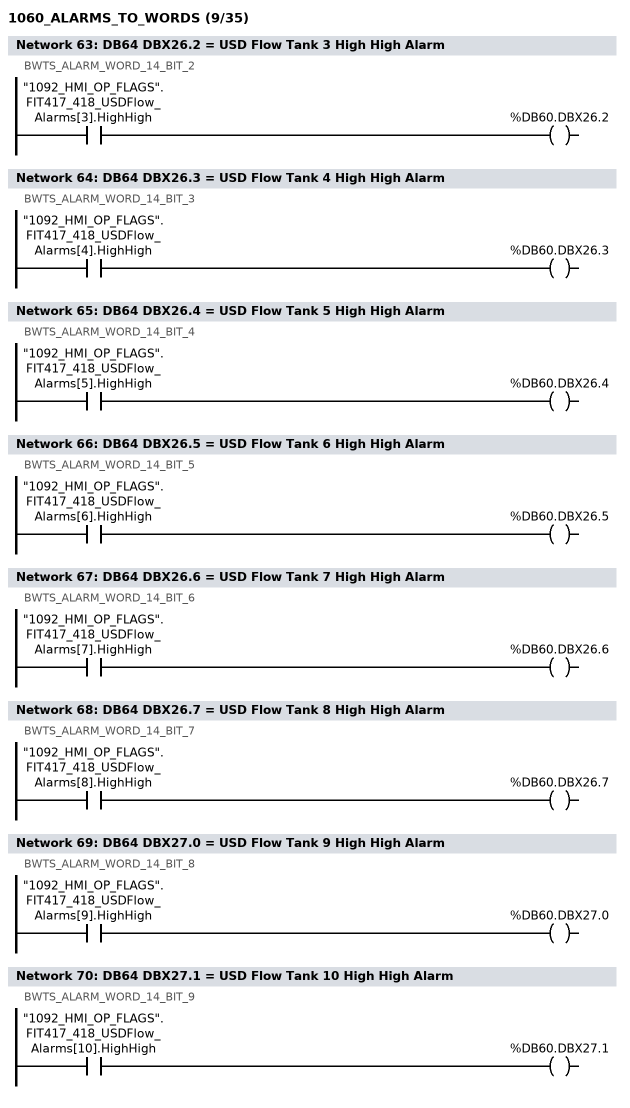
   RUNG wire#powerrail
      Contact( "1092_HMI_OP_FLAGS".FIT417_418_USDFlow_Alarms[3].HighHigh )
      Coil( %DB60.DBX26.2 )
   END_RUNG
   // the same network as SCL:
   %DB60.DBX26.2 := "1092_HMI_OP_FLAGS".FIT417_418_USDFlow_Alarms[3].HighHigh;
END_REGION

REGION Network 64: DB64 DBX26.3 = USD Flow Tank 4 High High Alarm
   // BWTS_ALARM_WORD_14_BIT_3
   RUNG wire#powerrail
      Contact( "1092_HMI_OP_FLAGS".FIT417_418_USDFlow_Alarms[4].HighHigh )
      Coil( %DB60.DBX26.3 )
   END_RUNG
   // the same network as SCL:
   %DB60.DBX26.3 := "1092_HMI_OP_FLAGS".FIT417_418_USDFlow_Alarms[4].HighHigh;
END_REGION

REGION Network 65: DB64 DBX26.4 = USD Flow Tank 5 High High Alarm
   // BWTS_ALARM_WORD_14_BIT_4
   RUNG wire#powerrail
      Contact( "1092_HMI_OP_FLAGS".FIT417_418_USDFlow_Alarms[5].HighHigh )
      Coil( %DB60.DBX26.4 )
   END_RUNG
   // the same network as SCL:
   %DB60.DBX26.4 := "1092_HMI_OP_FLAGS".FIT417_418_USDFlow_Alarms[5].HighHigh;
END_REGION

REGION Network 66: DB64 DBX26.5 = USD Flow Tank 6 High High Alarm
   // BWTS_ALARM_WORD_14_BIT_5
   RUNG wire#powerrail
      Contact( "1092_HMI_OP_FLAGS".FIT417_418_USDFlow_Alarms[6].HighHigh )
      Coil( %DB60.DBX26.5 )
   END_RUNG
   // the same network as SCL:
   %DB60.DBX26.5 := "1092_HMI_OP_FLAGS".FIT417_418_USDFlow_Alarms[6].HighHigh;
END_REGION

REGION Network 67: DB64 DBX26.6 = USD Flow Tank 7 High High Alarm
   // BWTS_ALARM_WORD_14_BIT_6
   RUNG wire#powerrail
      Contact( "1092_HMI_OP_FLAGS".FIT417_418_USDFlow_Alarms[7].HighHigh )
      Coil( %DB60.DBX26.6 )
   END_RUNG
   // the same network as SCL:
   %DB60.DBX26.6 := "1092_HMI_OP_FLAGS".FIT417_418_USDFlow_Alarms[7].HighHigh;
END_REGION

REGION Network 68: DB64 DBX26.7 = USD Flow Tank 8 High High Alarm
   // BWTS_ALARM_WORD_14_BIT_7
   RUNG wire#powerrail
      Contact( "1092_HMI_OP_FLAGS".FIT417_418_USDFlow_Alarms[8].HighHigh )
      Coil( %DB60.DBX26.7 )
   END_RUNG
   // the same network as SCL:
   %DB60.DBX26.7 := "1092_HMI_OP_FLAGS".FIT417_418_USDFlow_Alarms[8].HighHigh;
END_REGION

REGION Network 69: DB64 DBX27.0 = USD Flow Tank 9 High High Alarm
   // BWTS_ALARM_WORD_14_BIT_8
   RUNG wire#powerrail
      Contact( "1092_HMI_OP_FLAGS".FIT417_418_USDFlow_Alarms[9].HighHigh )
      Coil( %DB60.DBX27.0 )
   END_RUNG
   // the same network as SCL:
   %DB60.DBX27.0 := "1092_HMI_OP_FLAGS".FIT417_418_USDFlow_Alarms[9].HighHigh;
END_REGION

REGION Network 70: DB64 DBX27.1 = USD Flow Tank 10 High High Alarm
   // BWTS_ALARM_WORD_14_BIT_9
   RUNG wire#powerrail
      Contact( "1092_HMI_OP_FLAGS".FIT417_418_USDFlow_Alarms[10].HighHigh )
      Coil( %DB60.DBX27.1 )
   END_RUNG
   // the same network as SCL:
   %DB60.DBX27.1 := "1092_HMI_OP_FLAGS".FIT417_418_USDFlow_Alarms[10].HighHigh;
END_REGION

REGION Network 71: DB64 DBX27.2 = USD Flow Tank 11 High High Alarm
   // BWTS_ALARM_WORD_14_BIT_10
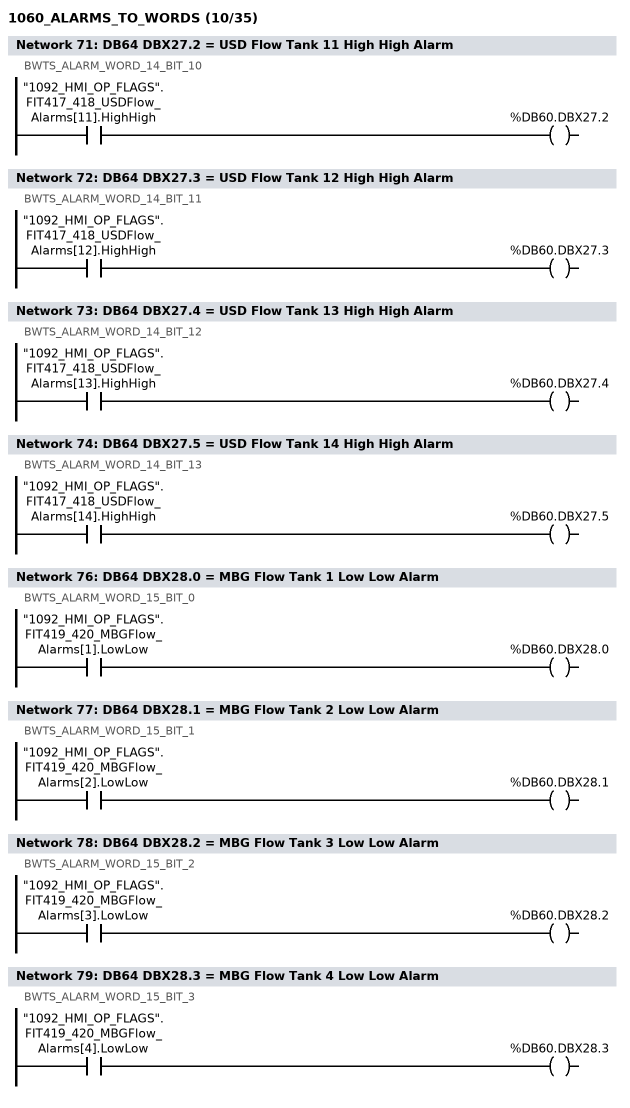
   RUNG wire#powerrail
      Contact( "1092_HMI_OP_FLAGS".FIT417_418_USDFlow_Alarms[11].HighHigh )
      Coil( %DB60.DBX27.2 )
   END_RUNG
   // the same network as SCL:
   %DB60.DBX27.2 := "1092_HMI_OP_FLAGS".FIT417_418_USDFlow_Alarms[11].HighHigh;
END_REGION

REGION Network 72: DB64 DBX27.3 = USD Flow Tank 12 High High Alarm
   // BWTS_ALARM_WORD_14_BIT_11
   RUNG wire#powerrail
      Contact( "1092_HMI_OP_FLAGS".FIT417_418_USDFlow_Alarms[12].HighHigh )
      Coil( %DB60.DBX27.3 )
   END_RUNG
   // the same network as SCL:
   %DB60.DBX27.3 := "1092_HMI_OP_FLAGS".FIT417_418_USDFlow_Alarms[12].HighHigh;
END_REGION

REGION Network 73: DB64 DBX27.4 = USD Flow Tank 13 High High Alarm
   // BWTS_ALARM_WORD_14_BIT_12
   RUNG wire#powerrail
      Contact( "1092_HMI_OP_FLAGS".FIT417_418_USDFlow_Alarms[13].HighHigh )
      Coil( %DB60.DBX27.4 )
   END_RUNG
   // the same network as SCL:
   %DB60.DBX27.4 := "1092_HMI_OP_FLAGS".FIT417_418_USDFlow_Alarms[13].HighHigh;
END_REGION

REGION Network 74: DB64 DBX27.5 = USD Flow Tank 14 High High Alarm
   // BWTS_ALARM_WORD_14_BIT_13
   RUNG wire#powerrail
      Contact( "1092_HMI_OP_FLAGS".FIT417_418_USDFlow_Alarms[14].HighHigh )
      Coil( %DB60.DBX27.5 )
   END_RUNG
   // the same network as SCL:
   %DB60.DBX27.5 := "1092_HMI_OP_FLAGS".FIT417_418_USDFlow_Alarms[14].HighHigh;
END_REGION

REGION Network 76: DB64 DBX28.0 = MBG Flow Tank 1 Low Low Alarm
   // BWTS_ALARM_WORD_15_BIT_0
   RUNG wire#powerrail
      Contact( "1092_HMI_OP_FLAGS".FIT419_420_MBGFlow_Alarms[1].LowLow )
      Coil( %DB60.DBX28.0 )
   END_RUNG
   // the same network as SCL:
   %DB60.DBX28.0 := "1092_HMI_OP_FLAGS".FIT419_420_MBGFlow_Alarms[1].LowLow;
END_REGION

REGION Network 77: DB64 DBX28.1 = MBG Flow Tank 2 Low Low Alarm
   // BWTS_ALARM_WORD_15_BIT_1
   RUNG wire#powerrail
      Contact( "1092_HMI_OP_FLAGS".FIT419_420_MBGFlow_Alarms[2].LowLow )
      Coil( %DB60.DBX28.1 )
   END_RUNG
   // the same network as SCL:
   %DB60.DBX28.1 := "1092_HMI_OP_FLAGS".FIT419_420_MBGFlow_Alarms[2].LowLow;
END_REGION

REGION Network 78: DB64 DBX28.2 = MBG Flow Tank 3 Low Low Alarm
   // BWTS_ALARM_WORD_15_BIT_2
   RUNG wire#powerrail
      Contact( "1092_HMI_OP_FLAGS".FIT419_420_MBGFlow_Alarms[3].LowLow )
      Coil( %DB60.DBX28.2 )
   END_RUNG
   // the same network as SCL:
   %DB60.DBX28.2 := "1092_HMI_OP_FLAGS".FIT419_420_MBGFlow_Alarms[3].LowLow;
END_REGION

REGION Network 79: DB64 DBX28.3 = MBG Flow Tank 4 Low Low Alarm
   // BWTS_ALARM_WORD_15_BIT_3
   RUNG wire#powerrail
      Contact( "1092_HMI_OP_FLAGS".FIT419_420_MBGFlow_Alarms[4].LowLow )
      Coil( %DB60.DBX28.3 )
   END_RUNG
   // the same network as SCL:
   %DB60.DBX28.3 := "1092_HMI_OP_FLAGS".FIT419_420_MBGFlow_Alarms[4].LowLow;
END_REGION

REGION Network 80: DB64 DBX28.4 = MBG Flow Tank 5 Low Low Alarm
   // BWTS_ALARM_WORD_15_BIT_4
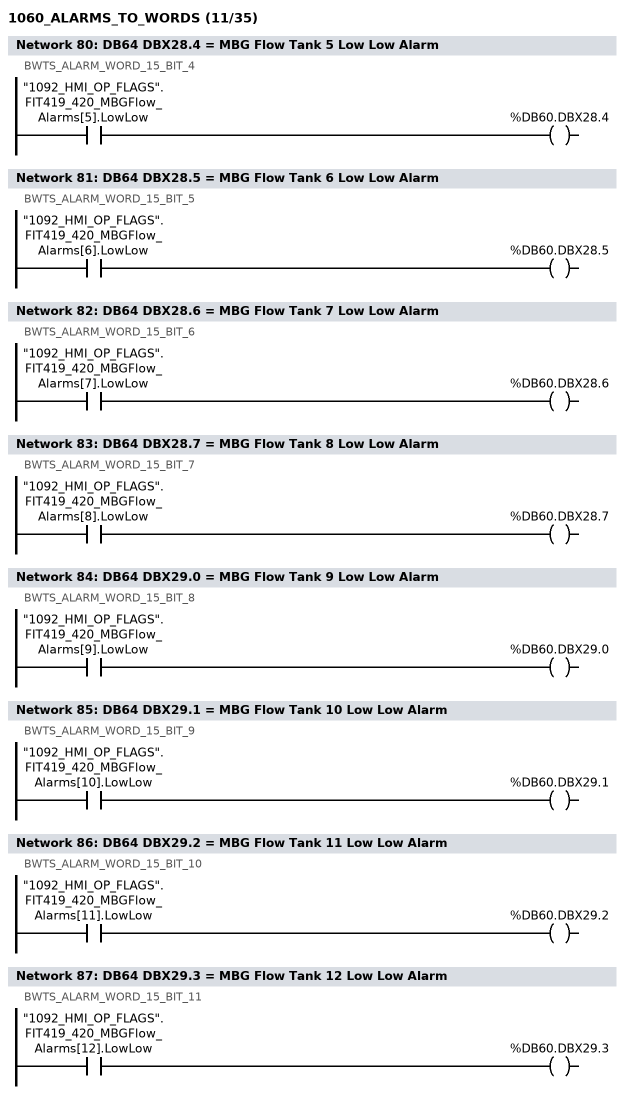
   RUNG wire#powerrail
      Contact( "1092_HMI_OP_FLAGS".FIT419_420_MBGFlow_Alarms[5].LowLow )
      Coil( %DB60.DBX28.4 )
   END_RUNG
   // the same network as SCL:
   %DB60.DBX28.4 := "1092_HMI_OP_FLAGS".FIT419_420_MBGFlow_Alarms[5].LowLow;
END_REGION

REGION Network 81: DB64 DBX28.5 = MBG Flow Tank 6 Low Low Alarm
   // BWTS_ALARM_WORD_15_BIT_5
   RUNG wire#powerrail
      Contact( "1092_HMI_OP_FLAGS".FIT419_420_MBGFlow_Alarms[6].LowLow )
      Coil( %DB60.DBX28.5 )
   END_RUNG
   // the same network as SCL:
   %DB60.DBX28.5 := "1092_HMI_OP_FLAGS".FIT419_420_MBGFlow_Alarms[6].LowLow;
END_REGION

REGION Network 82: DB64 DBX28.6 = MBG Flow Tank 7 Low Low Alarm
   // BWTS_ALARM_WORD_15_BIT_6
   RUNG wire#powerrail
      Contact( "1092_HMI_OP_FLAGS".FIT419_420_MBGFlow_Alarms[7].LowLow )
      Coil( %DB60.DBX28.6 )
   END_RUNG
   // the same network as SCL:
   %DB60.DBX28.6 := "1092_HMI_OP_FLAGS".FIT419_420_MBGFlow_Alarms[7].LowLow;
END_REGION

REGION Network 83: DB64 DBX28.7 = MBG Flow Tank 8 Low Low Alarm
   // BWTS_ALARM_WORD_15_BIT_7
   RUNG wire#powerrail
      Contact( "1092_HMI_OP_FLAGS".FIT419_420_MBGFlow_Alarms[8].LowLow )
      Coil( %DB60.DBX28.7 )
   END_RUNG
   // the same network as SCL:
   %DB60.DBX28.7 := "1092_HMI_OP_FLAGS".FIT419_420_MBGFlow_Alarms[8].LowLow;
END_REGION

REGION Network 84: DB64 DBX29.0 = MBG Flow Tank 9 Low Low Alarm
   // BWTS_ALARM_WORD_15_BIT_8
   RUNG wire#powerrail
      Contact( "1092_HMI_OP_FLAGS".FIT419_420_MBGFlow_Alarms[9].LowLow )
      Coil( %DB60.DBX29.0 )
   END_RUNG
   // the same network as SCL:
   %DB60.DBX29.0 := "1092_HMI_OP_FLAGS".FIT419_420_MBGFlow_Alarms[9].LowLow;
END_REGION

REGION Network 85: DB64 DBX29.1 = MBG Flow Tank 10 Low Low Alarm
   // BWTS_ALARM_WORD_15_BIT_9
   RUNG wire#powerrail
      Contact( "1092_HMI_OP_FLAGS".FIT419_420_MBGFlow_Alarms[10].LowLow )
      Coil( %DB60.DBX29.1 )
   END_RUNG
   // the same network as SCL:
   %DB60.DBX29.1 := "1092_HMI_OP_FLAGS".FIT419_420_MBGFlow_Alarms[10].LowLow;
END_REGION

REGION Network 86: DB64 DBX29.2 = MBG Flow Tank 11 Low Low Alarm
   // BWTS_ALARM_WORD_15_BIT_10
   RUNG wire#powerrail
      Contact( "1092_HMI_OP_FLAGS".FIT419_420_MBGFlow_Alarms[11].LowLow )
      Coil( %DB60.DBX29.2 )
   END_RUNG
   // the same network as SCL:
   %DB60.DBX29.2 := "1092_HMI_OP_FLAGS".FIT419_420_MBGFlow_Alarms[11].LowLow;
END_REGION

REGION Network 87: DB64 DBX29.3 = MBG Flow Tank 12 Low Low Alarm
   // BWTS_ALARM_WORD_15_BIT_11
   RUNG wire#powerrail
      Contact( "1092_HMI_OP_FLAGS".FIT419_420_MBGFlow_Alarms[12].LowLow )
      Coil( %DB60.DBX29.3 )
   END_RUNG
   // the same network as SCL:
   %DB60.DBX29.3 := "1092_HMI_OP_FLAGS".FIT419_420_MBGFlow_Alarms[12].LowLow;
END_REGION

REGION Network 88: DB64 DBX29.4 = MBG Flow Tank 13 Low Low Alarm
   // BWTS_ALARM_WORD_15_BIT_12
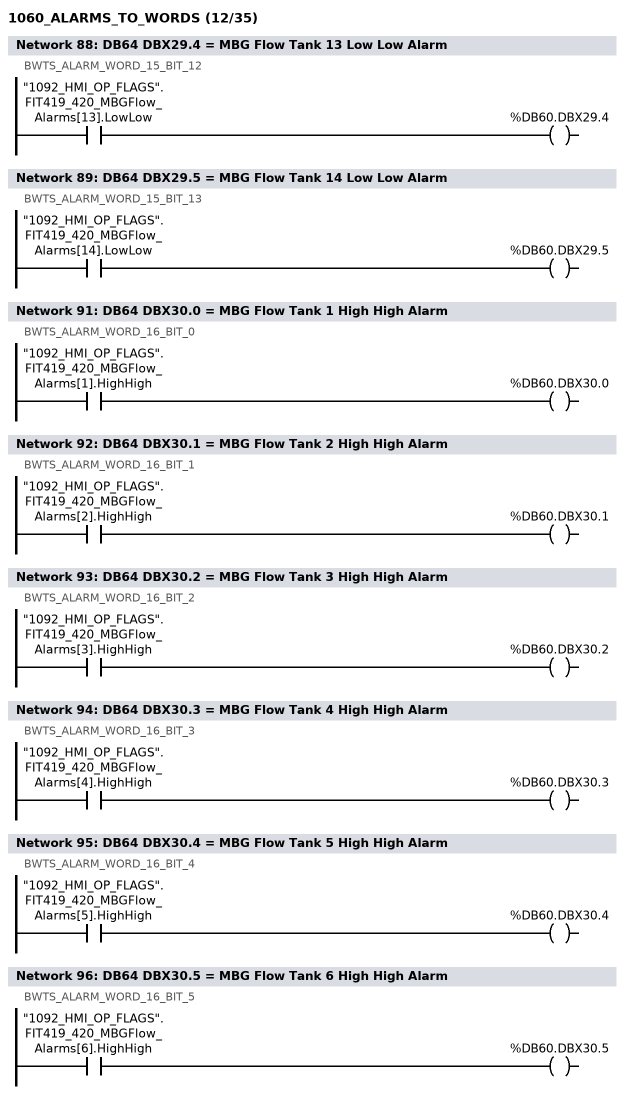
   RUNG wire#powerrail
      Contact( "1092_HMI_OP_FLAGS".FIT419_420_MBGFlow_Alarms[13].LowLow )
      Coil( %DB60.DBX29.4 )
   END_RUNG
   // the same network as SCL:
   %DB60.DBX29.4 := "1092_HMI_OP_FLAGS".FIT419_420_MBGFlow_Alarms[13].LowLow;
END_REGION

REGION Network 89: DB64 DBX29.5 = MBG Flow Tank 14 Low Low Alarm
   // BWTS_ALARM_WORD_15_BIT_13
   RUNG wire#powerrail
      Contact( "1092_HMI_OP_FLAGS".FIT419_420_MBGFlow_Alarms[14].LowLow )
      Coil( %DB60.DBX29.5 )
   END_RUNG
   // the same network as SCL:
   %DB60.DBX29.5 := "1092_HMI_OP_FLAGS".FIT419_420_MBGFlow_Alarms[14].LowLow;
END_REGION

REGION Network 91: DB64 DBX30.0 = MBG Flow Tank 1 High High Alarm
   // BWTS_ALARM_WORD_16_BIT_0
   RUNG wire#powerrail
      Contact( "1092_HMI_OP_FLAGS".FIT419_420_MBGFlow_Alarms[1].HighHigh )
      Coil( %DB60.DBX30.0 )
   END_RUNG
   // the same network as SCL:
   %DB60.DBX30.0 := "1092_HMI_OP_FLAGS".FIT419_420_MBGFlow_Alarms[1].HighHigh;
END_REGION

REGION Network 92: DB64 DBX30.1 = MBG Flow Tank 2 High High Alarm
   // BWTS_ALARM_WORD_16_BIT_1
   RUNG wire#powerrail
      Contact( "1092_HMI_OP_FLAGS".FIT419_420_MBGFlow_Alarms[2].HighHigh )
      Coil( %DB60.DBX30.1 )
   END_RUNG
   // the same network as SCL:
   %DB60.DBX30.1 := "1092_HMI_OP_FLAGS".FIT419_420_MBGFlow_Alarms[2].HighHigh;
END_REGION

REGION Network 93: DB64 DBX30.2 = MBG Flow Tank 3 High High Alarm
   // BWTS_ALARM_WORD_16_BIT_2
   RUNG wire#powerrail
      Contact( "1092_HMI_OP_FLAGS".FIT419_420_MBGFlow_Alarms[3].HighHigh )
      Coil( %DB60.DBX30.2 )
   END_RUNG
   // the same network as SCL:
   %DB60.DBX30.2 := "1092_HMI_OP_FLAGS".FIT419_420_MBGFlow_Alarms[3].HighHigh;
END_REGION

REGION Network 94: DB64 DBX30.3 = MBG Flow Tank 4 High High Alarm
   // BWTS_ALARM_WORD_16_BIT_3
   RUNG wire#powerrail
      Contact( "1092_HMI_OP_FLAGS".FIT419_420_MBGFlow_Alarms[4].HighHigh )
      Coil( %DB60.DBX30.3 )
   END_RUNG
   // the same network as SCL:
   %DB60.DBX30.3 := "1092_HMI_OP_FLAGS".FIT419_420_MBGFlow_Alarms[4].HighHigh;
END_REGION

REGION Network 95: DB64 DBX30.4 = MBG Flow Tank 5 High High Alarm
   // BWTS_ALARM_WORD_16_BIT_4
   RUNG wire#powerrail
      Contact( "1092_HMI_OP_FLAGS".FIT419_420_MBGFlow_Alarms[5].HighHigh )
      Coil( %DB60.DBX30.4 )
   END_RUNG
   // the same network as SCL:
   %DB60.DBX30.4 := "1092_HMI_OP_FLAGS".FIT419_420_MBGFlow_Alarms[5].HighHigh;
END_REGION

REGION Network 96: DB64 DBX30.5 = MBG Flow Tank 6 High High Alarm
   // BWTS_ALARM_WORD_16_BIT_5
   RUNG wire#powerrail
      Contact( "1092_HMI_OP_FLAGS".FIT419_420_MBGFlow_Alarms[6].HighHigh )
      Coil( %DB60.DBX30.5 )
   END_RUNG
   // the same network as SCL:
   %DB60.DBX30.5 := "1092_HMI_OP_FLAGS".FIT419_420_MBGFlow_Alarms[6].HighHigh;
END_REGION

REGION Network 97: DB64 DBX30.6 = MBG Flow Tank 7 High High Alarm
   // BWTS_ALARM_WORD_16_BIT_6
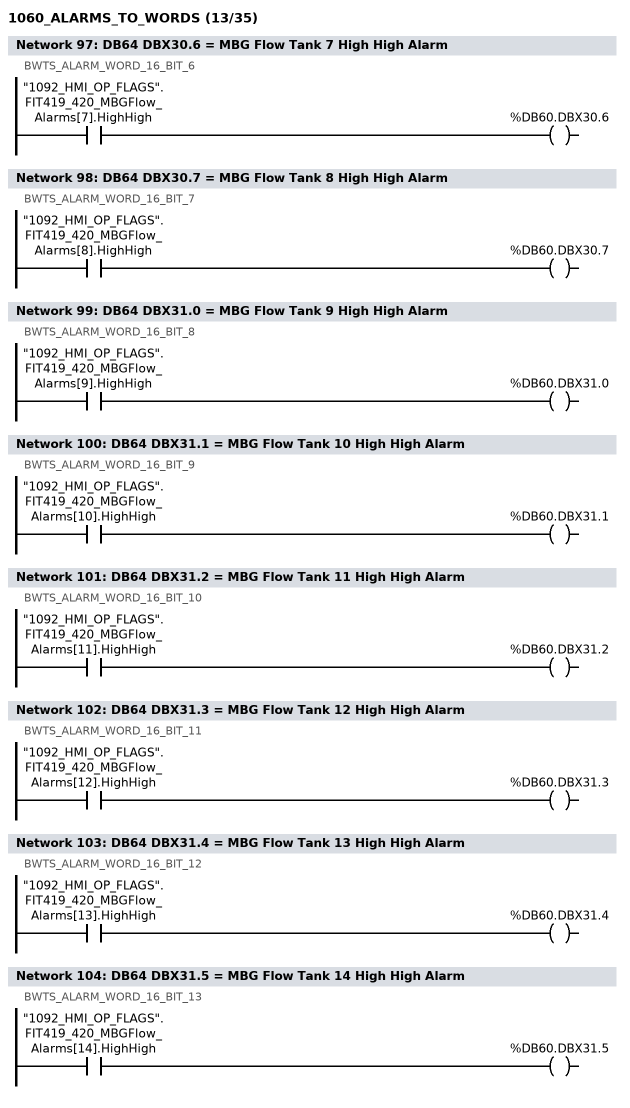
   RUNG wire#powerrail
      Contact( "1092_HMI_OP_FLAGS".FIT419_420_MBGFlow_Alarms[7].HighHigh )
      Coil( %DB60.DBX30.6 )
   END_RUNG
   // the same network as SCL:
   %DB60.DBX30.6 := "1092_HMI_OP_FLAGS".FIT419_420_MBGFlow_Alarms[7].HighHigh;
END_REGION

REGION Network 98: DB64 DBX30.7 = MBG Flow Tank 8 High High Alarm
   // BWTS_ALARM_WORD_16_BIT_7
   RUNG wire#powerrail
      Contact( "1092_HMI_OP_FLAGS".FIT419_420_MBGFlow_Alarms[8].HighHigh )
      Coil( %DB60.DBX30.7 )
   END_RUNG
   // the same network as SCL:
   %DB60.DBX30.7 := "1092_HMI_OP_FLAGS".FIT419_420_MBGFlow_Alarms[8].HighHigh;
END_REGION

REGION Network 99: DB64 DBX31.0 = MBG Flow Tank 9 High High Alarm
   // BWTS_ALARM_WORD_16_BIT_8
   RUNG wire#powerrail
      Contact( "1092_HMI_OP_FLAGS".FIT419_420_MBGFlow_Alarms[9].HighHigh )
      Coil( %DB60.DBX31.0 )
   END_RUNG
   // the same network as SCL:
   %DB60.DBX31.0 := "1092_HMI_OP_FLAGS".FIT419_420_MBGFlow_Alarms[9].HighHigh;
END_REGION

REGION Network 100: DB64 DBX31.1 = MBG Flow Tank 10 High High Alarm
   // BWTS_ALARM_WORD_16_BIT_9
   RUNG wire#powerrail
      Contact( "1092_HMI_OP_FLAGS".FIT419_420_MBGFlow_Alarms[10].HighHigh )
      Coil( %DB60.DBX31.1 )
   END_RUNG
   // the same network as SCL:
   %DB60.DBX31.1 := "1092_HMI_OP_FLAGS".FIT419_420_MBGFlow_Alarms[10].HighHigh;
END_REGION

REGION Network 101: DB64 DBX31.2 = MBG Flow Tank 11 High High Alarm
   // BWTS_ALARM_WORD_16_BIT_10
   RUNG wire#powerrail
      Contact( "1092_HMI_OP_FLAGS".FIT419_420_MBGFlow_Alarms[11].HighHigh )
      Coil( %DB60.DBX31.2 )
   END_RUNG
   // the same network as SCL:
   %DB60.DBX31.2 := "1092_HMI_OP_FLAGS".FIT419_420_MBGFlow_Alarms[11].HighHigh;
END_REGION

REGION Network 102: DB64 DBX31.3 = MBG Flow Tank 12 High High Alarm
   // BWTS_ALARM_WORD_16_BIT_11
   RUNG wire#powerrail
      Contact( "1092_HMI_OP_FLAGS".FIT419_420_MBGFlow_Alarms[12].HighHigh )
      Coil( %DB60.DBX31.3 )
   END_RUNG
   // the same network as SCL:
   %DB60.DBX31.3 := "1092_HMI_OP_FLAGS".FIT419_420_MBGFlow_Alarms[12].HighHigh;
END_REGION

REGION Network 103: DB64 DBX31.4 = MBG Flow Tank 13 High High Alarm
   // BWTS_ALARM_WORD_16_BIT_12
   RUNG wire#powerrail
      Contact( "1092_HMI_OP_FLAGS".FIT419_420_MBGFlow_Alarms[13].HighHigh )
      Coil( %DB60.DBX31.4 )
   END_RUNG
   // the same network as SCL:
   %DB60.DBX31.4 := "1092_HMI_OP_FLAGS".FIT419_420_MBGFlow_Alarms[13].HighHigh;
END_REGION

REGION Network 104: DB64 DBX31.5 = MBG Flow Tank 14 High High Alarm
   // BWTS_ALARM_WORD_16_BIT_13
   RUNG wire#powerrail
      Contact( "1092_HMI_OP_FLAGS".FIT419_420_MBGFlow_Alarms[14].HighHigh )
      Coil( %DB60.DBX31.5 )
   END_RUNG
   // the same network as SCL:
   %DB60.DBX31.5 := "1092_HMI_OP_FLAGS".FIT419_420_MBGFlow_Alarms[14].HighHigh;
END_REGION

REGION Network 106: DB64 DBX32.0 = BWT Level Tank 1 Low Alarm
   // BWTS_ALARM_WORD_17_BIT_0
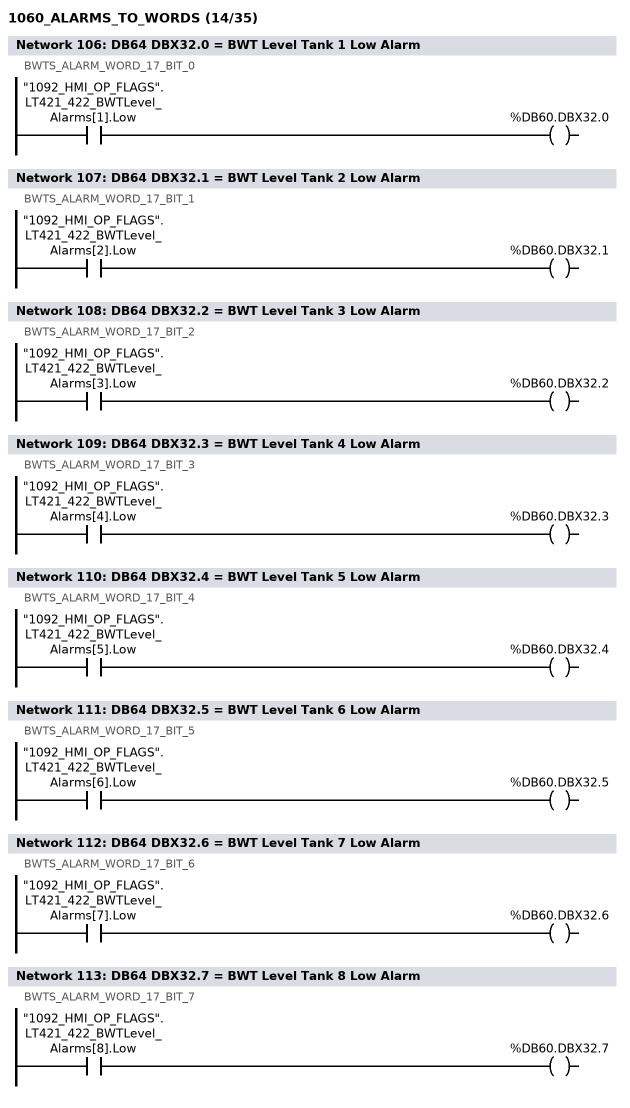
   RUNG wire#powerrail
      Contact( "1092_HMI_OP_FLAGS".LT421_422_BWTLevel_Alarms[1].Low )
      Coil( %DB60.DBX32.0 )
   END_RUNG
   // the same network as SCL:
   %DB60.DBX32.0 := "1092_HMI_OP_FLAGS".LT421_422_BWTLevel_Alarms[1].Low;
END_REGION

REGION Network 107: DB64 DBX32.1 = BWT Level Tank 2 Low Alarm
   // BWTS_ALARM_WORD_17_BIT_1
   RUNG wire#powerrail
      Contact( "1092_HMI_OP_FLAGS".LT421_422_BWTLevel_Alarms[2].Low )
      Coil( %DB60.DBX32.1 )
   END_RUNG
   // the same network as SCL:
   %DB60.DBX32.1 := "1092_HMI_OP_FLAGS".LT421_422_BWTLevel_Alarms[2].Low;
END_REGION

REGION Network 108: DB64 DBX32.2 = BWT Level Tank 3 Low Alarm
   // BWTS_ALARM_WORD_17_BIT_2
   RUNG wire#powerrail
      Contact( "1092_HMI_OP_FLAGS".LT421_422_BWTLevel_Alarms[3].Low )
      Coil( %DB60.DBX32.2 )
   END_RUNG
   // the same network as SCL:
   %DB60.DBX32.2 := "1092_HMI_OP_FLAGS".LT421_422_BWTLevel_Alarms[3].Low;
END_REGION

REGION Network 109: DB64 DBX32.3 = BWT Level Tank 4 Low Alarm
   // BWTS_ALARM_WORD_17_BIT_3
   RUNG wire#powerrail
      Contact( "1092_HMI_OP_FLAGS".LT421_422_BWTLevel_Alarms[4].Low )
      Coil( %DB60.DBX32.3 )
   END_RUNG
   // the same network as SCL:
   %DB60.DBX32.3 := "1092_HMI_OP_FLAGS".LT421_422_BWTLevel_Alarms[4].Low;
END_REGION

REGION Network 110: DB64 DBX32.4 = BWT Level Tank 5 Low Alarm
   // BWTS_ALARM_WORD_17_BIT_4
   RUNG wire#powerrail
      Contact( "1092_HMI_OP_FLAGS".LT421_422_BWTLevel_Alarms[5].Low )
      Coil( %DB60.DBX32.4 )
   END_RUNG
   // the same network as SCL:
   %DB60.DBX32.4 := "1092_HMI_OP_FLAGS".LT421_422_BWTLevel_Alarms[5].Low;
END_REGION

REGION Network 111: DB64 DBX32.5 = BWT Level Tank 6 Low Alarm
   // BWTS_ALARM_WORD_17_BIT_5
   RUNG wire#powerrail
      Contact( "1092_HMI_OP_FLAGS".LT421_422_BWTLevel_Alarms[6].Low )
      Coil( %DB60.DBX32.5 )
   END_RUNG
   // the same network as SCL:
   %DB60.DBX32.5 := "1092_HMI_OP_FLAGS".LT421_422_BWTLevel_Alarms[6].Low;
END_REGION

REGION Network 112: DB64 DBX32.6 = BWT Level Tank 7 Low Alarm
   // BWTS_ALARM_WORD_17_BIT_6
   RUNG wire#powerrail
      Contact( "1092_HMI_OP_FLAGS".LT421_422_BWTLevel_Alarms[7].Low )
      Coil( %DB60.DBX32.6 )
   END_RUNG
   // the same network as SCL:
   %DB60.DBX32.6 := "1092_HMI_OP_FLAGS".LT421_422_BWTLevel_Alarms[7].Low;
END_REGION

REGION Network 113: DB64 DBX32.7 = BWT Level Tank 8 Low Alarm
   // BWTS_ALARM_WORD_17_BIT_7
   RUNG wire#powerrail
      Contact( "1092_HMI_OP_FLAGS".LT421_422_BWTLevel_Alarms[8].Low )
      Coil( %DB60.DBX32.7 )
   END_RUNG
   // the same network as SCL:
   %DB60.DBX32.7 := "1092_HMI_OP_FLAGS".LT421_422_BWTLevel_Alarms[8].Low;
END_REGION

REGION Network 114: DB64 DBX33.0 = BWT Level Tank 9 Low Alarm
   // BWTS_ALARM_WORD_17_BIT_8
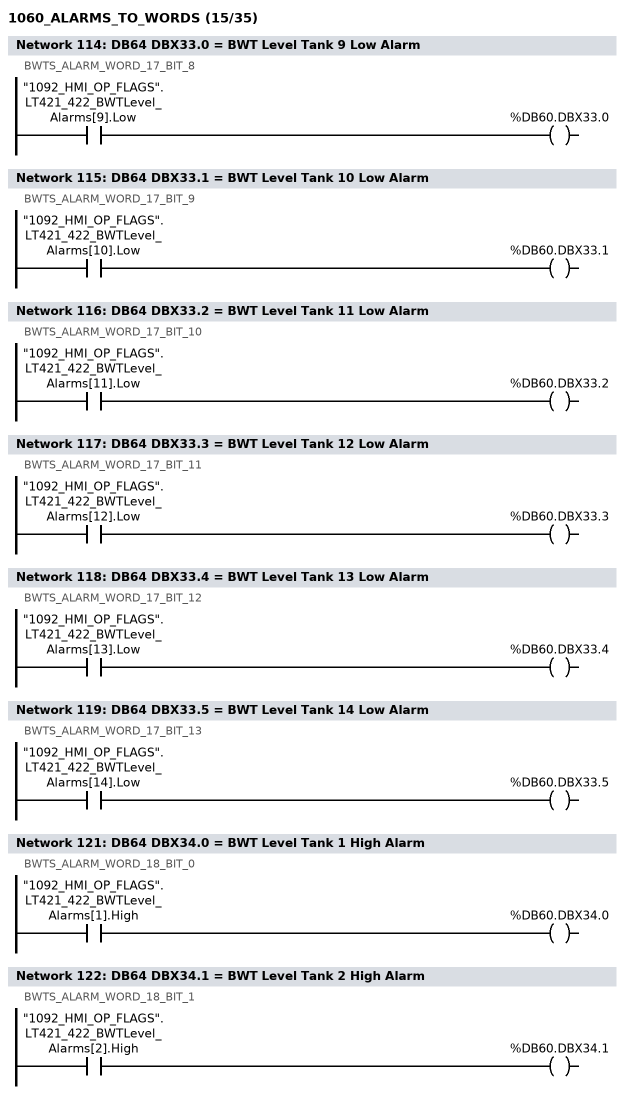
   RUNG wire#powerrail
      Contact( "1092_HMI_OP_FLAGS".LT421_422_BWTLevel_Alarms[9].Low )
      Coil( %DB60.DBX33.0 )
   END_RUNG
   // the same network as SCL:
   %DB60.DBX33.0 := "1092_HMI_OP_FLAGS".LT421_422_BWTLevel_Alarms[9].Low;
END_REGION

REGION Network 115: DB64 DBX33.1 = BWT Level Tank 10 Low Alarm
   // BWTS_ALARM_WORD_17_BIT_9
   RUNG wire#powerrail
      Contact( "1092_HMI_OP_FLAGS".LT421_422_BWTLevel_Alarms[10].Low )
      Coil( %DB60.DBX33.1 )
   END_RUNG
   // the same network as SCL:
   %DB60.DBX33.1 := "1092_HMI_OP_FLAGS".LT421_422_BWTLevel_Alarms[10].Low;
END_REGION

REGION Network 116: DB64 DBX33.2 = BWT Level Tank 11 Low Alarm
   // BWTS_ALARM_WORD_17_BIT_10
   RUNG wire#powerrail
      Contact( "1092_HMI_OP_FLAGS".LT421_422_BWTLevel_Alarms[11].Low )
      Coil( %DB60.DBX33.2 )
   END_RUNG
   // the same network as SCL:
   %DB60.DBX33.2 := "1092_HMI_OP_FLAGS".LT421_422_BWTLevel_Alarms[11].Low;
END_REGION

REGION Network 117: DB64 DBX33.3 = BWT Level Tank 12 Low Alarm
   // BWTS_ALARM_WORD_17_BIT_11
   RUNG wire#powerrail
      Contact( "1092_HMI_OP_FLAGS".LT421_422_BWTLevel_Alarms[12].Low )
      Coil( %DB60.DBX33.3 )
   END_RUNG
   // the same network as SCL:
   %DB60.DBX33.3 := "1092_HMI_OP_FLAGS".LT421_422_BWTLevel_Alarms[12].Low;
END_REGION

REGION Network 118: DB64 DBX33.4 = BWT Level Tank 13 Low Alarm
   // BWTS_ALARM_WORD_17_BIT_12
   RUNG wire#powerrail
      Contact( "1092_HMI_OP_FLAGS".LT421_422_BWTLevel_Alarms[13].Low )
      Coil( %DB60.DBX33.4 )
   END_RUNG
   // the same network as SCL:
   %DB60.DBX33.4 := "1092_HMI_OP_FLAGS".LT421_422_BWTLevel_Alarms[13].Low;
END_REGION

REGION Network 119: DB64 DBX33.5 = BWT Level Tank 14 Low Alarm
   // BWTS_ALARM_WORD_17_BIT_13
   RUNG wire#powerrail
      Contact( "1092_HMI_OP_FLAGS".LT421_422_BWTLevel_Alarms[14].Low )
      Coil( %DB60.DBX33.5 )
   END_RUNG
   // the same network as SCL:
   %DB60.DBX33.5 := "1092_HMI_OP_FLAGS".LT421_422_BWTLevel_Alarms[14].Low;
END_REGION

REGION Network 121: DB64 DBX34.0 = BWT Level Tank 1 High Alarm
   // BWTS_ALARM_WORD_18_BIT_0
   RUNG wire#powerrail
      Contact( "1092_HMI_OP_FLAGS".LT421_422_BWTLevel_Alarms[1].High )
      Coil( %DB60.DBX34.0 )
   END_RUNG
   // the same network as SCL:
   %DB60.DBX34.0 := "1092_HMI_OP_FLAGS".LT421_422_BWTLevel_Alarms[1].High;
END_REGION

REGION Network 122: DB64 DBX34.1 = BWT Level Tank 2 High Alarm
   // BWTS_ALARM_WORD_18_BIT_1
   RUNG wire#powerrail
      Contact( "1092_HMI_OP_FLAGS".LT421_422_BWTLevel_Alarms[2].High )
      Coil( %DB60.DBX34.1 )
   END_RUNG
   // the same network as SCL:
   %DB60.DBX34.1 := "1092_HMI_OP_FLAGS".LT421_422_BWTLevel_Alarms[2].High;
END_REGION

REGION Network 123: DB64 DBX34.2 = BWT Level Tank 3 High Alarm
   // BWTS_ALARM_WORD_18_BIT_2
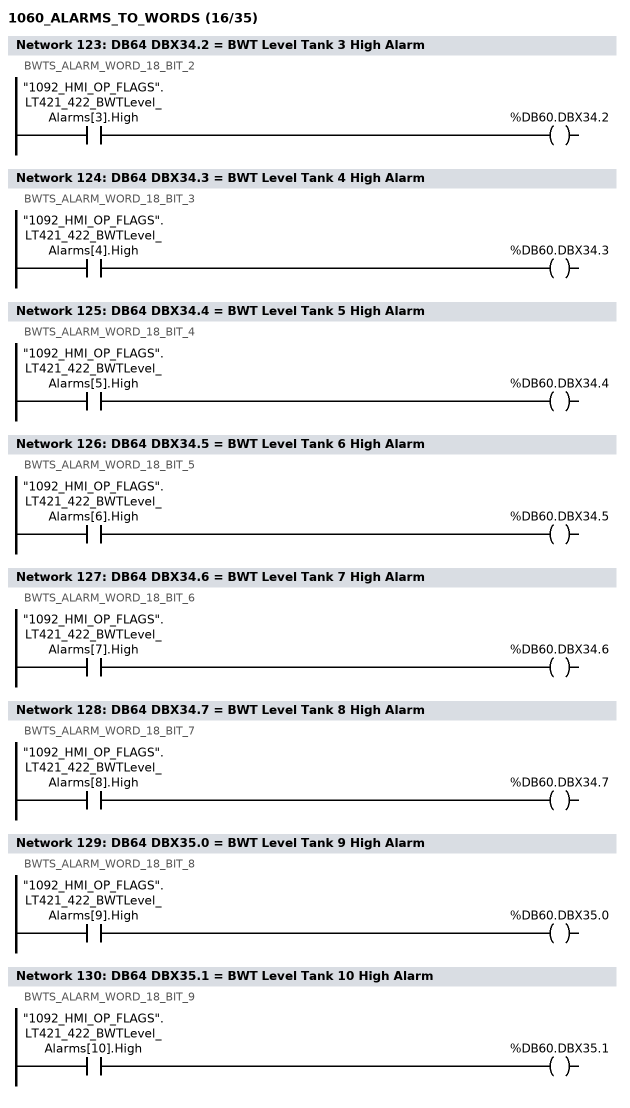
   RUNG wire#powerrail
      Contact( "1092_HMI_OP_FLAGS".LT421_422_BWTLevel_Alarms[3].High )
      Coil( %DB60.DBX34.2 )
   END_RUNG
   // the same network as SCL:
   %DB60.DBX34.2 := "1092_HMI_OP_FLAGS".LT421_422_BWTLevel_Alarms[3].High;
END_REGION

REGION Network 124: DB64 DBX34.3 = BWT Level Tank 4 High Alarm
   // BWTS_ALARM_WORD_18_BIT_3
   RUNG wire#powerrail
      Contact( "1092_HMI_OP_FLAGS".LT421_422_BWTLevel_Alarms[4].High )
      Coil( %DB60.DBX34.3 )
   END_RUNG
   // the same network as SCL:
   %DB60.DBX34.3 := "1092_HMI_OP_FLAGS".LT421_422_BWTLevel_Alarms[4].High;
END_REGION

REGION Network 125: DB64 DBX34.4 = BWT Level Tank 5 High Alarm
   // BWTS_ALARM_WORD_18_BIT_4
   RUNG wire#powerrail
      Contact( "1092_HMI_OP_FLAGS".LT421_422_BWTLevel_Alarms[5].High )
      Coil( %DB60.DBX34.4 )
   END_RUNG
   // the same network as SCL:
   %DB60.DBX34.4 := "1092_HMI_OP_FLAGS".LT421_422_BWTLevel_Alarms[5].High;
END_REGION

REGION Network 126: DB64 DBX34.5 = BWT Level Tank 6 High Alarm
   // BWTS_ALARM_WORD_18_BIT_5
   RUNG wire#powerrail
      Contact( "1092_HMI_OP_FLAGS".LT421_422_BWTLevel_Alarms[6].High )
      Coil( %DB60.DBX34.5 )
   END_RUNG
   // the same network as SCL:
   %DB60.DBX34.5 := "1092_HMI_OP_FLAGS".LT421_422_BWTLevel_Alarms[6].High;
END_REGION

REGION Network 127: DB64 DBX34.6 = BWT Level Tank 7 High Alarm
   // BWTS_ALARM_WORD_18_BIT_6
   RUNG wire#powerrail
      Contact( "1092_HMI_OP_FLAGS".LT421_422_BWTLevel_Alarms[7].High )
      Coil( %DB60.DBX34.6 )
   END_RUNG
   // the same network as SCL:
   %DB60.DBX34.6 := "1092_HMI_OP_FLAGS".LT421_422_BWTLevel_Alarms[7].High;
END_REGION

REGION Network 128: DB64 DBX34.7 = BWT Level Tank 8 High Alarm
   // BWTS_ALARM_WORD_18_BIT_7
   RUNG wire#powerrail
      Contact( "1092_HMI_OP_FLAGS".LT421_422_BWTLevel_Alarms[8].High )
      Coil( %DB60.DBX34.7 )
   END_RUNG
   // the same network as SCL:
   %DB60.DBX34.7 := "1092_HMI_OP_FLAGS".LT421_422_BWTLevel_Alarms[8].High;
END_REGION

REGION Network 129: DB64 DBX35.0 = BWT Level Tank 9 High Alarm
   // BWTS_ALARM_WORD_18_BIT_8
   RUNG wire#powerrail
      Contact( "1092_HMI_OP_FLAGS".LT421_422_BWTLevel_Alarms[9].High )
      Coil( %DB60.DBX35.0 )
   END_RUNG
   // the same network as SCL:
   %DB60.DBX35.0 := "1092_HMI_OP_FLAGS".LT421_422_BWTLevel_Alarms[9].High;
END_REGION

REGION Network 130: DB64 DBX35.1 = BWT Level Tank 10 High Alarm
   // BWTS_ALARM_WORD_18_BIT_9
   RUNG wire#powerrail
      Contact( "1092_HMI_OP_FLAGS".LT421_422_BWTLevel_Alarms[10].High )
      Coil( %DB60.DBX35.1 )
   END_RUNG
   // the same network as SCL:
   %DB60.DBX35.1 := "1092_HMI_OP_FLAGS".LT421_422_BWTLevel_Alarms[10].High;
END_REGION

REGION Network 131: DB64 DBX35.2 = BWT Level Tank 11 High Alarm
   // BWTS_ALARM_WORD_18_BIT_10
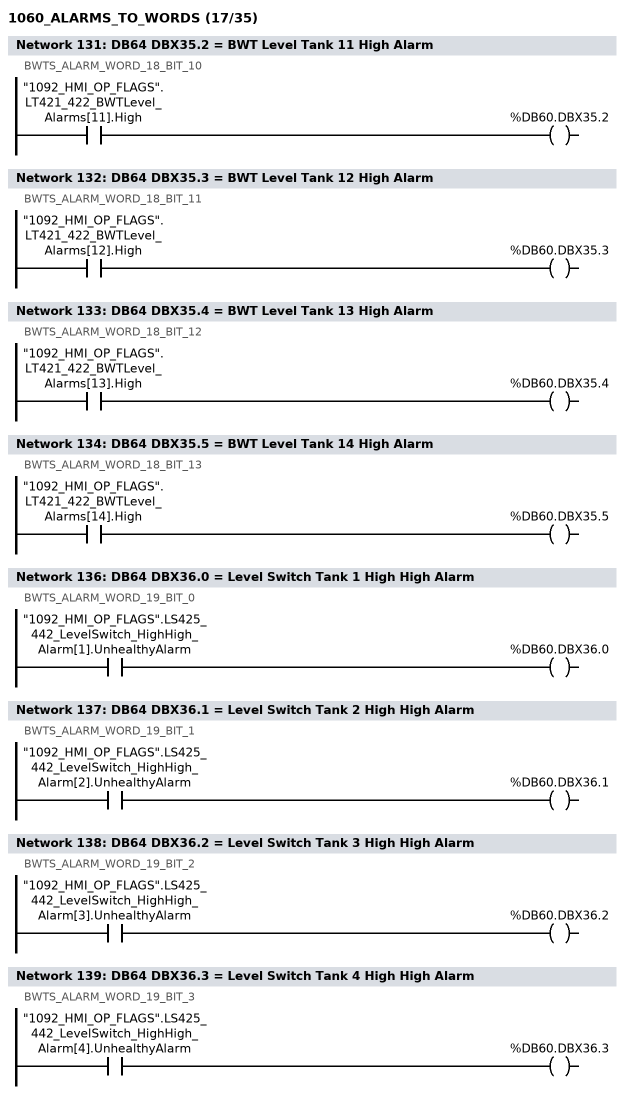
   RUNG wire#powerrail
      Contact( "1092_HMI_OP_FLAGS".LT421_422_BWTLevel_Alarms[11].High )
      Coil( %DB60.DBX35.2 )
   END_RUNG
   // the same network as SCL:
   %DB60.DBX35.2 := "1092_HMI_OP_FLAGS".LT421_422_BWTLevel_Alarms[11].High;
END_REGION

REGION Network 132: DB64 DBX35.3 = BWT Level Tank 12 High Alarm
   // BWTS_ALARM_WORD_18_BIT_11
   RUNG wire#powerrail
      Contact( "1092_HMI_OP_FLAGS".LT421_422_BWTLevel_Alarms[12].High )
      Coil( %DB60.DBX35.3 )
   END_RUNG
   // the same network as SCL:
   %DB60.DBX35.3 := "1092_HMI_OP_FLAGS".LT421_422_BWTLevel_Alarms[12].High;
END_REGION

REGION Network 133: DB64 DBX35.4 = BWT Level Tank 13 High Alarm
   // BWTS_ALARM_WORD_18_BIT_12
   RUNG wire#powerrail
      Contact( "1092_HMI_OP_FLAGS".LT421_422_BWTLevel_Alarms[13].High )
      Coil( %DB60.DBX35.4 )
   END_RUNG
   // the same network as SCL:
   %DB60.DBX35.4 := "1092_HMI_OP_FLAGS".LT421_422_BWTLevel_Alarms[13].High;
END_REGION

REGION Network 134: DB64 DBX35.5 = BWT Level Tank 14 High Alarm
   // BWTS_ALARM_WORD_18_BIT_13
   RUNG wire#powerrail
      Contact( "1092_HMI_OP_FLAGS".LT421_422_BWTLevel_Alarms[14].High )
      Coil( %DB60.DBX35.5 )
   END_RUNG
   // the same network as SCL:
   %DB60.DBX35.5 := "1092_HMI_OP_FLAGS".LT421_422_BWTLevel_Alarms[14].High;
END_REGION

REGION Network 136: DB64 DBX36.0 = Level Switch Tank 1 High High Alarm
   // BWTS_ALARM_WORD_19_BIT_0
   RUNG wire#powerrail
      Contact( "1092_HMI_OP_FLAGS".LS425_442_LevelSwitch_HighHigh_Alarm[1].UnhealthyAlarm )
      Coil( %DB60.DBX36.0 )
   END_RUNG
   // the same network as SCL:
   %DB60.DBX36.0 := "1092_HMI_OP_FLAGS".LS425_442_LevelSwitch_HighHigh_Alarm[1].UnhealthyAlarm;
END_REGION

REGION Network 137: DB64 DBX36.1 = Level Switch Tank 2 High High Alarm
   // BWTS_ALARM_WORD_19_BIT_1
   RUNG wire#powerrail
      Contact( "1092_HMI_OP_FLAGS".LS425_442_LevelSwitch_HighHigh_Alarm[2].UnhealthyAlarm )
      Coil( %DB60.DBX36.1 )
   END_RUNG
   // the same network as SCL:
   %DB60.DBX36.1 := "1092_HMI_OP_FLAGS".LS425_442_LevelSwitch_HighHigh_Alarm[2].UnhealthyAlarm;
END_REGION

REGION Network 138: DB64 DBX36.2 = Level Switch Tank 3 High High Alarm
   // BWTS_ALARM_WORD_19_BIT_2
   RUNG wire#powerrail
      Contact( "1092_HMI_OP_FLAGS".LS425_442_LevelSwitch_HighHigh_Alarm[3].UnhealthyAlarm )
      Coil( %DB60.DBX36.2 )
   END_RUNG
   // the same network as SCL:
   %DB60.DBX36.2 := "1092_HMI_OP_FLAGS".LS425_442_LevelSwitch_HighHigh_Alarm[3].UnhealthyAlarm;
END_REGION

REGION Network 139: DB64 DBX36.3 = Level Switch Tank 4 High High Alarm
   // BWTS_ALARM_WORD_19_BIT_3
   RUNG wire#powerrail
      Contact( "1092_HMI_OP_FLAGS".LS425_442_LevelSwitch_HighHigh_Alarm[4].UnhealthyAlarm )
      Coil( %DB60.DBX36.3 )
   END_RUNG
   // the same network as SCL:
   %DB60.DBX36.3 := "1092_HMI_OP_FLAGS".LS425_442_LevelSwitch_HighHigh_Alarm[4].UnhealthyAlarm;
END_REGION

REGION Network 140: DB64 DBX36.4 = Level Switch Tank 5 High High Alarm
   // BWTS_ALARM_WORD_19_BIT_4
